(* Logix 5000 project; controller _GigaDiscovery vendor 1 type 14 code 244 rev 35.11; software revision 35.03; part 18 of 23 *)
(* tags used below, declared in another part *)
   Home_Timer : TIMER;
   Timer2 : TIMER;
   DC_Field_Motor_7 : UDT_CROUT;   // DC Field Motor 7 Gondola Contactor -Q16101E -Q16103E
   DC_Field_Pylon_Motors : UDT_CROUT;   // DC Field Pylon Motors Contactor -Q10101E -Q10103E
   FeedBack_Drives_Contactors : BOOL;
   Gate_Entry_Unlock_Selector : BOOL;   // -S30701F
   Gate_Exit_Unlock_Selector : BOOL;   // -S30705F
   Gate_Operator_Unlock_Selector : BOOL;   // -S30707F
   Gondola_Drive_Enable : UDT_CROUT;   // Gondola Drive Ch1-Ch2 Start Enable Contactors -Q16105E -Q16107E
   Gondola_Standstill_from_inertia : BOOL;
   I_Fbk_Platform_Main_Valve : UDT_DCS;   // Feedback Platform Main Valve -B21902I
   I_Fire_Interface : UDT_DCM;   // Page 44
   I_Gate_ENTER_G01_Closed : UDT_DCM;   // GATE ENTER (G01) -B25204I
   I_Gate_EXIT_G05_Closed : UDT_DCM;   // GATE EXIT (G05) -B25304I
   I_Gate_OPERATOR_Closed : UDT_DCM;   // GATE 4 OPERATOR RFID SENSOR - MOP -B25404J
   I_Gates_Closed : UDT_DCM;   // Gate Closed RFID series -B24802J
   I_GMB_RCC1_Temperature_OK : BOOL;   // +GMB_RCC1 Temperature OK -S40103E
   I_Gondola_Home_Position : BOOL;   // Gondola Home Position -B40002I -B40007I
   I_Gondola_Home_Position_Sensor_1 : UDT_DCM;   // Home Sensor Speed Check -B40002I
   I_Gondola_Home_Position_Sensor_2 : UDT_DCM;   // Home Sensor Speed Check -B40007I
   I_Platform_Closed : UDT_DCM;   // Platform Closed RFID Series -B22501J... -B22807J -B22801B
   I_Platform_Line_Min_Pressure_Switch : BOOL;   // Platform Line Minimum Pressure Switch -S21511B
   I_Platform_Line_Unlock_Pressure_Switch : BOOL;   // Unlock Platform Line Pressure Switch -S22006B
   I_Platform_Opened : UDT_DCM;   // Platform Opened RFID Series -Q23801J -Q23807J
   I_Platform_Pressure_on_Close_Circuit : BOOL;   // Platform Maximum Closing Pressure -S21510B
   I_Platform_Pressure_on_Open_Circuit : BOOL;   // Platform Maximum Opening Pressure -S21507B
   I_Pylon_Home_Ch1 : UDT_DCM;   // Home position Pylon Ch1 -B26002I
   I_Pylon_Home_Ch2 : UDT_DCM;   // Home position Pylon Ch2 -B26007I
   I_Pylon_Overlimit_Right : UDT_DCS;   // Pylon Overlimit Switchs -A26510I
   I_RCC_GSA_Temperature_OK : BOOL;   // +RCC_GSA Temperature OK -S50110G
   I_RCC_GSB_Temperature_OK : BOOL;   // +RCC_GSB Temperature OK -S52110G
   I_RCC_GSC_Temperature_OK : BOOL;   // +RCC_GSC Temperature OK -S54110G
   I_RCC_GSD_Temperature_OK : BOOL;   // +RCC_GSD Temperature OK -S56110G
   I_RCC_GSE_Temperature_OK : BOOL;   // +RCC_GSE Temperature OK -S58110G
   I_RCC_GSF_Temperature_OK : BOOL;   // +RCC_GSF Temperature OK -S60110G
   I_RCC_GSG_Temperature_OK : BOOL;   // +RCC_GSG Temperature OK -S62110G
   I_RCC_GSH_Temperature_OK : BOOL;   // +RCC_GSH Temperature OK -S64110G
   I_RESTRAINTS_Close_Limit_Switch : BOOL;   // Main Valve Close Limit Switch -B40508I
   I_RESTRAINTS_Open_Limit_Switch : BOOL;   // Main Valve Open Limit Switch -B40504I
   O_RESTRAINTS_Main_Valve : BOOL;   // Main Valve -B40501I
   O_RESTRAINTS_MainValve : UDT_CROUT;   // Main Valve -B40501I
   ONP : DINT;   // Optional Not Present
   Platform_Fbk_Valv_Close : BOOL;   // Platform Close Main Valve Limit Switch -B21909I
   Platform_Fbk_Valv_Open : BOOL;   // Platform Open Main Valve Limit Switch -B21905I
   Power_On_Delay : BOOL;
   Pylon_Contactor_OFF : BOOL;
   Pylon_Home_Position : UDT_DCM;   // Home position Pylon -B26002I -B26007I
   Pylon_Start_Drive_1_2 : UDT_CROUT;   // Pylon Start Drive 1 - 2 Contactors -Q9002H -Q9004H -Q10202G
   Pylon_Start_Drive_3_4 : UDT_CROUT;   // Pylon Start Drive 3 - 4 Contactors -Q9005H -Q9007H -Q12202G
   Pylon_Start_Drive_5_6 : UDT_CROUT;   // Pylon Start Drive 5 - 6 Contactors -Q9009E -Q9011E4 -Q14202G -Q14202G
   Pylon_Stopped_At_Home : BOOL;   // 5s
   Reset_Pulse : BOOL;
   RESTRAINTS_MainValve_PressTest : Valve_2_pos_monostable;
   RESTRAINTS_Rack : LapBar_Racks[41];
   RESTRAINTS_Sector : LapBars_Sector[9];
   RESTRAINTS_Unlock_Valve_Pressure : BOOL;
   Valves_Pressure_Discrepancy : DINT;
(* S_Input, continued *)

ROUTINE _04_Platform   (* ladder *)
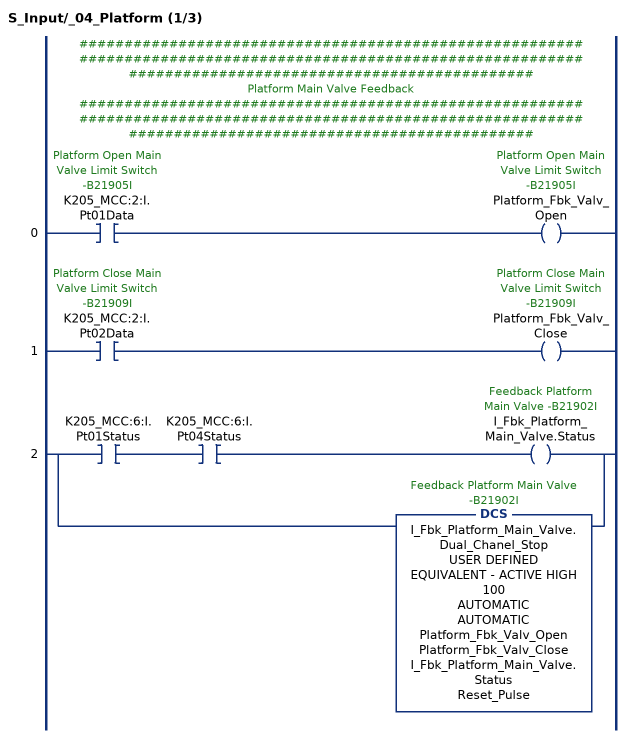
   // #############################################################################################################################################################
   // Platform Main Valve Feedback
   // #############################################################################################################################################################
   0: XIC(K205_MCC:2:I.Pt01Data)OTE(Platform_Fbk_Valv_Open);
   1: XIC(K205_MCC:2:I.Pt02Data)OTE(Platform_Fbk_Valv_Close);
   2: [XIC(K205_MCC:6:I.Pt01Status) XIC(K205_MCC:6:I.Pt04Status) OTE(I_Fbk_Platform_Main_Valve.Status) ,DCS(I_Fbk_Platform_Main_Valve.Dual_Chanel_Stop,USER DEFINED,EQUIVALENT - ACTIVE HIGH,100,AUTOMATIC,AUTOMATIC,Platform_Fbk_Valv_Open,Platform_Fbk_Valv_Close,I_Fbk_Platform_Main_Valve.Status,Reset_Pulse) ];
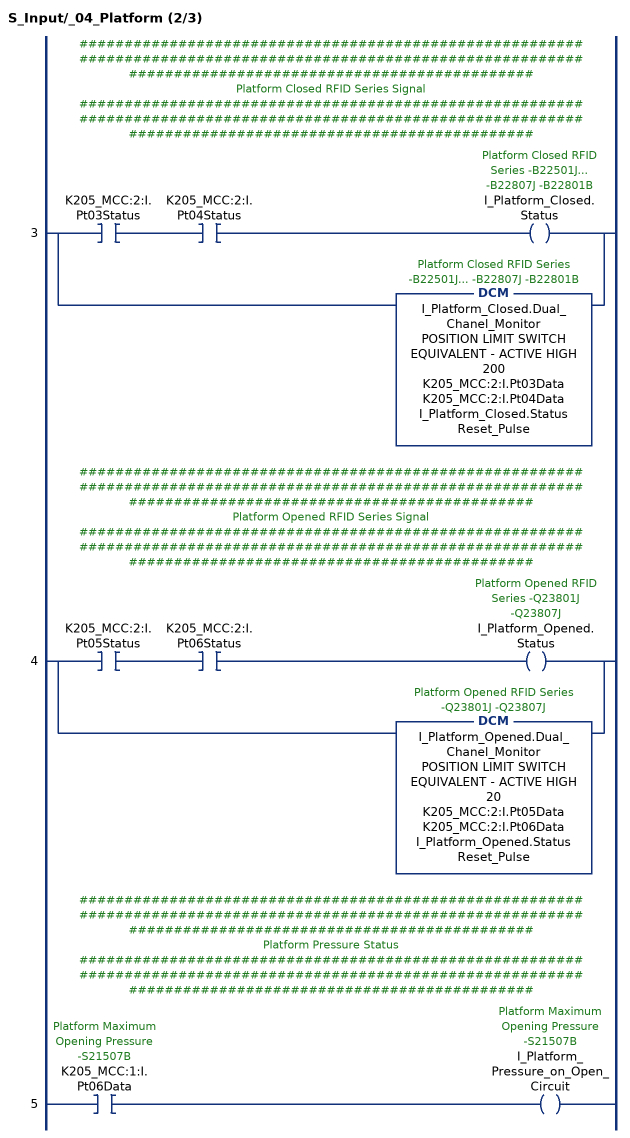
   // #############################################################################################################################################################
   // Platform Closed RFID Series Signal
   // #############################################################################################################################################################
   3: [XIC(K205_MCC:2:I.Pt03Status) XIC(K205_MCC:2:I.Pt04Status) OTE(I_Platform_Closed.Status) ,DCM(I_Platform_Closed.Dual_Chanel_Monitor,POSITION LIMIT SWITCH,EQUIVALENT - ACTIVE HIGH,200,K205_MCC:2:I.Pt03Data,K205_MCC:2:I.Pt04Data,I_Platform_Closed.Status,Reset_Pulse) ];
   // #############################################################################################################################################################
   // Platform Opened RFID Series Signal
   // #############################################################################################################################################################
   4: [XIC(K205_MCC:2:I.Pt05Status) XIC(K205_MCC:2:I.Pt06Status) OTE(I_Platform_Opened.Status) ,DCM(I_Platform_Opened.Dual_Chanel_Monitor,POSITION LIMIT SWITCH,EQUIVALENT - ACTIVE HIGH,20,K205_MCC:2:I.Pt05Data,K205_MCC:2:I.Pt06Data,I_Platform_Opened.Status,Reset_Pulse) ];
   // #############################################################################################################################################################
   // Platform Pressure Status
   // #############################################################################################################################################################
   5: XIC(K205_MCC:1:I.Pt06Data)OTE(I_Platform_Pressure_on_Open_Circuit);
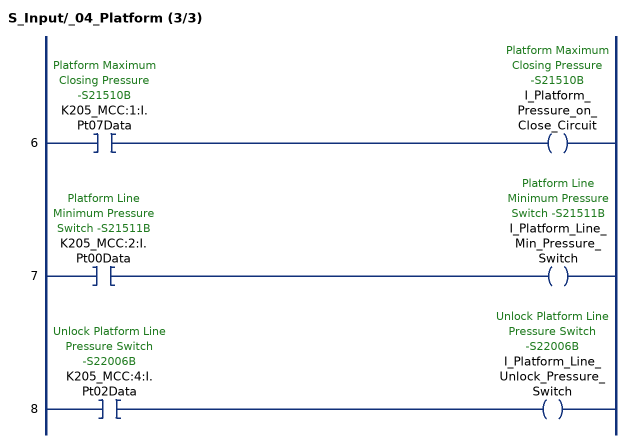
   6: XIC(K205_MCC:1:I.Pt07Data)OTE(I_Platform_Pressure_on_Close_Circuit);
   7: XIC(K205_MCC:2:I.Pt00Data)OTE(I_Platform_Line_Min_Pressure_Switch);
   8: XIC(K205_MCC:4:I.Pt02Data)OTE(I_Platform_Line_Unlock_Pressure_Switch);
END_ROUTINE

ROUTINE _05_Pylon   (* ladder *)
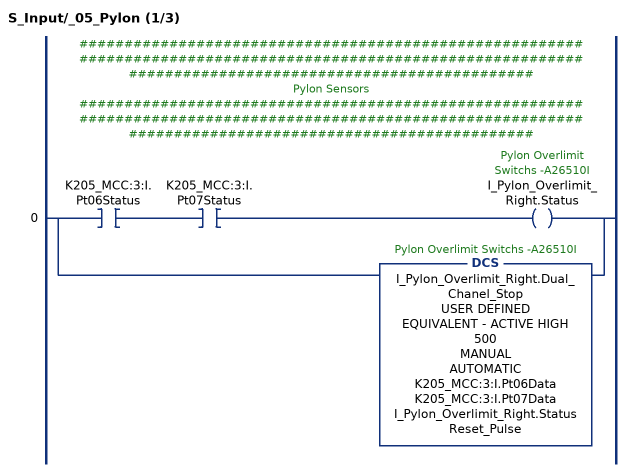
   // #############################################################################################################################################################
   // Pylon Sensors
   // #############################################################################################################################################################
   0: [XIC(K205_MCC:3:I.Pt06Status) XIC(K205_MCC:3:I.Pt07Status) OTE(I_Pylon_Overlimit_Right.Status) ,DCS(I_Pylon_Overlimit_Right.Dual_Chanel_Stop,USER DEFINED,EQUIVALENT - ACTIVE HIGH,500,MANUAL,AUTOMATIC,K205_MCC:3:I.Pt06Data,K205_MCC:3:I.Pt07Data,I_Pylon_Overlimit_Right.Status,Reset_Pulse) ];
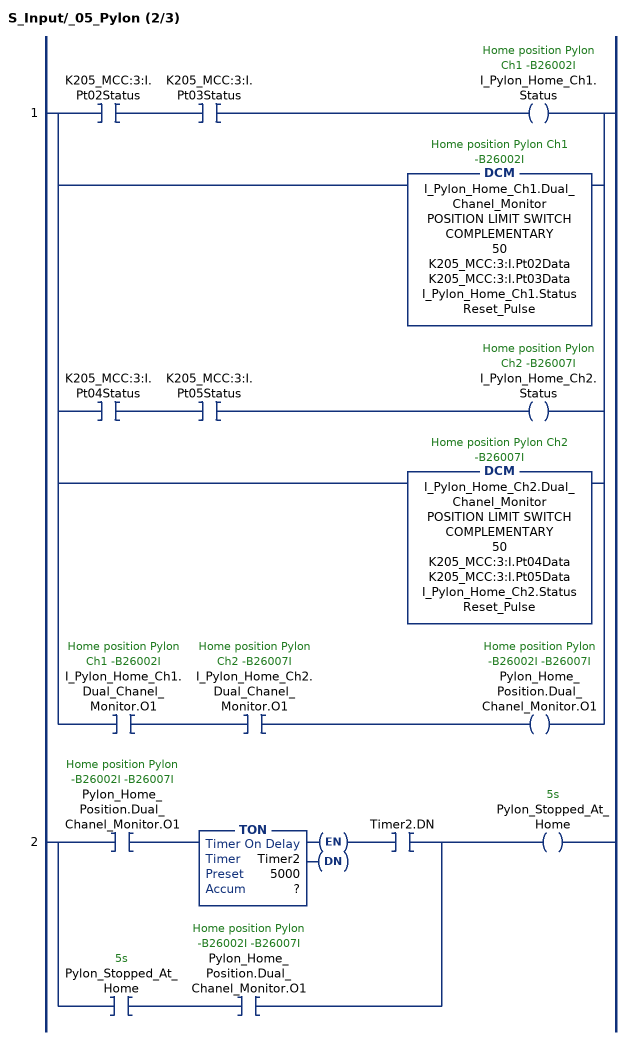
   1: [[XIC(K205_MCC:3:I.Pt02Status) XIC(K205_MCC:3:I.Pt03Status) OTE(I_Pylon_Home_Ch1.Status) ,DCM(I_Pylon_Home_Ch1.Dual_Chanel_Monitor,POSITION LIMIT SWITCH,COMPLEMENTARY,50,K205_MCC:3:I.Pt02Data,K205_MCC:3:I.Pt03Data,I_Pylon_Home_Ch1.Status,Reset_Pulse) ] ,[XIC(K205_MCC:3:I.Pt04Status) XIC(K205_MCC:3:I.Pt05Status) OTE(I_Pylon_Home_Ch2.Status) ,DCM(I_Pylon_Home_Ch2.Dual_Chanel_Monitor,POSITION LIMIT SWITCH,COMPLEMENTARY,50,K205_MCC:3:I.Pt04Data,K205_MCC:3:I.Pt05Data,I_Pylon_Home_Ch2.Status,Reset_Pulse) ] ,XIC(I_Pylon_Home_Ch1.Dual_Chanel_Monitor.O1) XIC(I_Pylon_Home_Ch2.Dual_Chanel_Monitor.O1) OTE(Pylon_Home_Position.Dual_Chanel_Monitor.O1) ];
   2: [XIC(Pylon_Home_Position.Dual_Chanel_Monitor.O1) TON(Timer2,?,?) XIC(Timer2.DN) ,XIC(Pylon_Stopped_At_Home) XIC(Pylon_Home_Position.Dual_Chanel_Monitor.O1) ]OTE(Pylon_Stopped_At_Home);
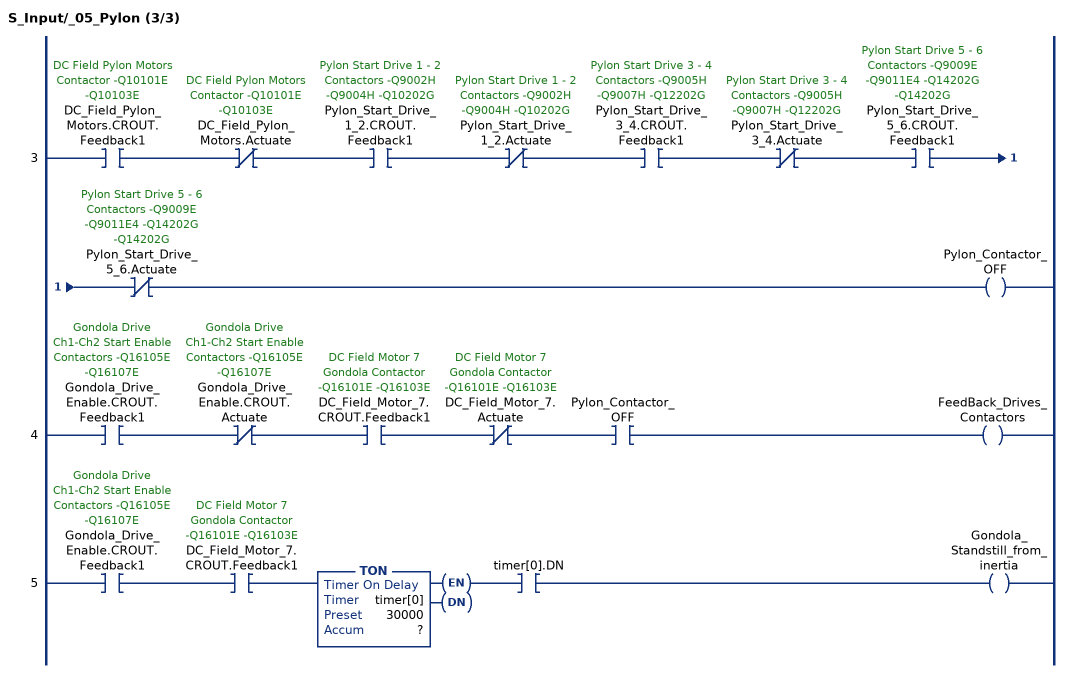
   3: XIC(DC_Field_Pylon_Motors.CROUT.Feedback1)XIO(DC_Field_Pylon_Motors.Actuate)XIC(Pylon_Start_Drive_1_2.CROUT.Feedback1)XIO(Pylon_Start_Drive_1_2.Actuate)XIC(Pylon_Start_Drive_3_4.CROUT.Feedback1)XIO(Pylon_Start_Drive_3_4.Actuate)XIC(Pylon_Start_Drive_5_6.CROUT.Feedback1)XIO(Pylon_Start_Drive_5_6.Actuate)OTE(Pylon_Contactor_OFF);
   4: XIC(Gondola_Drive_Enable.CROUT.Feedback1)XIO(Gondola_Drive_Enable.CROUT.Actuate)XIC(DC_Field_Motor_7.CROUT.Feedback1)XIO(DC_Field_Motor_7.Actuate)XIC(Pylon_Contactor_OFF)OTE(FeedBack_Drives_Contactors);
   5: XIC(Gondola_Drive_Enable.CROUT.Feedback1)XIC(DC_Field_Motor_7.CROUT.Feedback1)TON(timer[0],?,?)XIC(timer[0].DN)OTE(Gondola_Standstill_from_inertia);
END_ROUTINE

ROUTINE _06_RCC   (* ladder *)
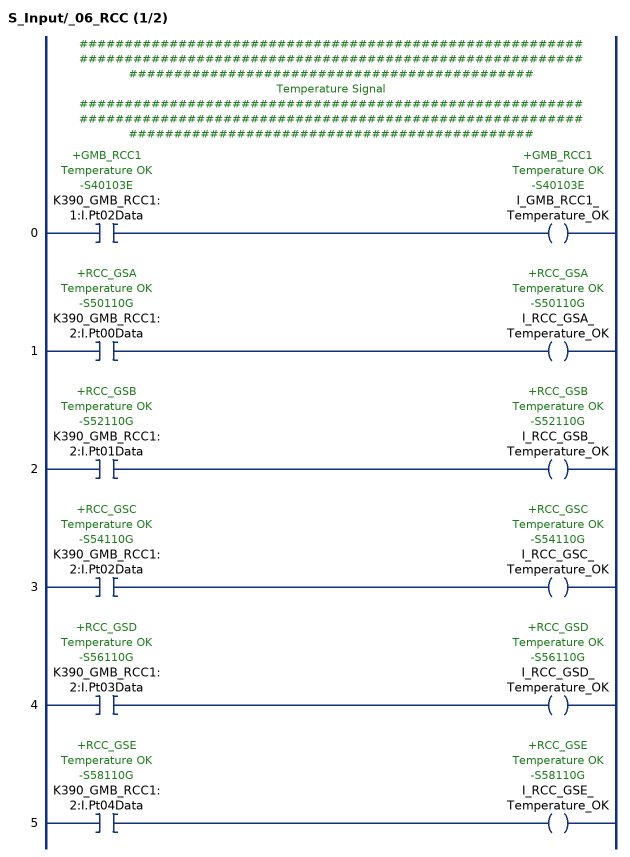
   // #############################################################################################################################################################
   //   Temperature Signal
   // #############################################################################################################################################################
   0: XIC(K390_GMB_RCC1:1:I.Pt02Data)OTE(I_GMB_RCC1_Temperature_OK);
   1: XIC(K390_GMB_RCC1:2:I.Pt00Data)OTE(I_RCC_GSA_Temperature_OK);
   2: XIC(K390_GMB_RCC1:2:I.Pt01Data)OTE(I_RCC_GSB_Temperature_OK);
   3: XIC(K390_GMB_RCC1:2:I.Pt02Data)OTE(I_RCC_GSC_Temperature_OK);
   4: XIC(K390_GMB_RCC1:2:I.Pt03Data)OTE(I_RCC_GSD_Temperature_OK);
   5: XIC(K390_GMB_RCC1:2:I.Pt04Data)OTE(I_RCC_GSE_Temperature_OK);
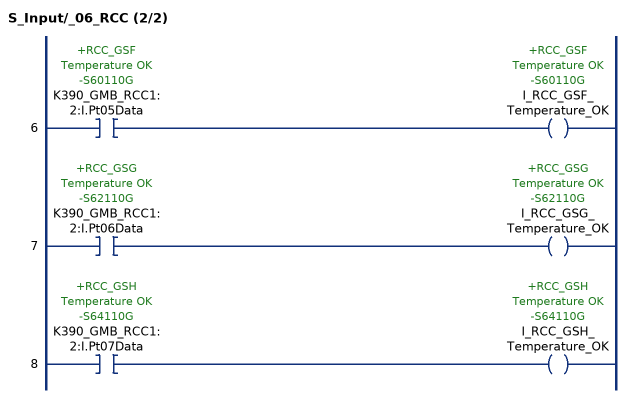
   6: XIC(K390_GMB_RCC1:2:I.Pt05Data)OTE(I_RCC_GSF_Temperature_OK);
   7: XIC(K390_GMB_RCC1:2:I.Pt06Data)OTE(I_RCC_GSG_Temperature_OK);
   8: XIC(K390_GMB_RCC1:2:I.Pt07Data)OTE(I_RCC_GSH_Temperature_OK);
END_ROUTINE

ROUTINE _07_Gate   (* ladder *)
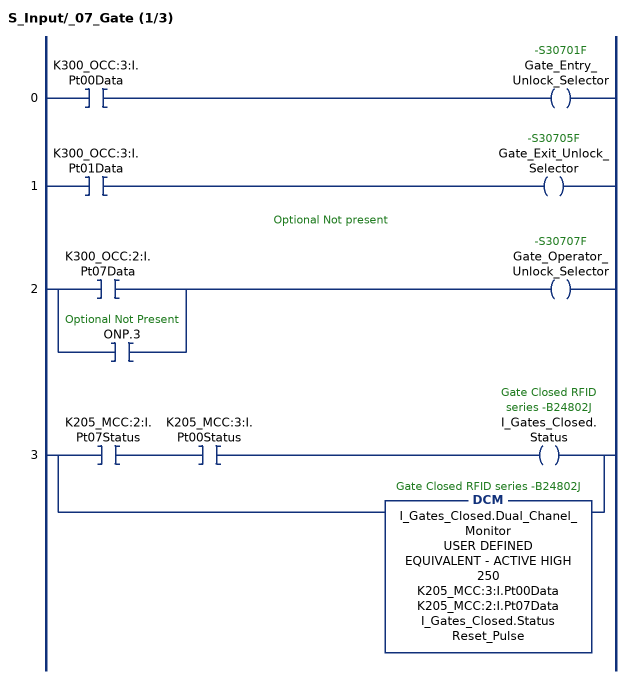
   0: XIC(K300_OCC:3:I.Pt00Data)OTE(Gate_Entry_Unlock_Selector);
   1: XIC(K300_OCC:3:I.Pt01Data)OTE(Gate_Exit_Unlock_Selector);
   // Optional Not present
   2: [XIC(K300_OCC:2:I.Pt07Data) ,XIC(ONP.3) ]OTE(Gate_Operator_Unlock_Selector);
   3: [XIC(K205_MCC:2:I.Pt07Status) XIC(K205_MCC:3:I.Pt00Status) OTE(I_Gates_Closed.Status) ,DCM(I_Gates_Closed.Dual_Chanel_Monitor,USER DEFINED,EQUIVALENT - ACTIVE HIGH,250,K205_MCC:3:I.Pt00Data,K205_MCC:2:I.Pt07Data,I_Gates_Closed.Status,Reset_Pulse) ];
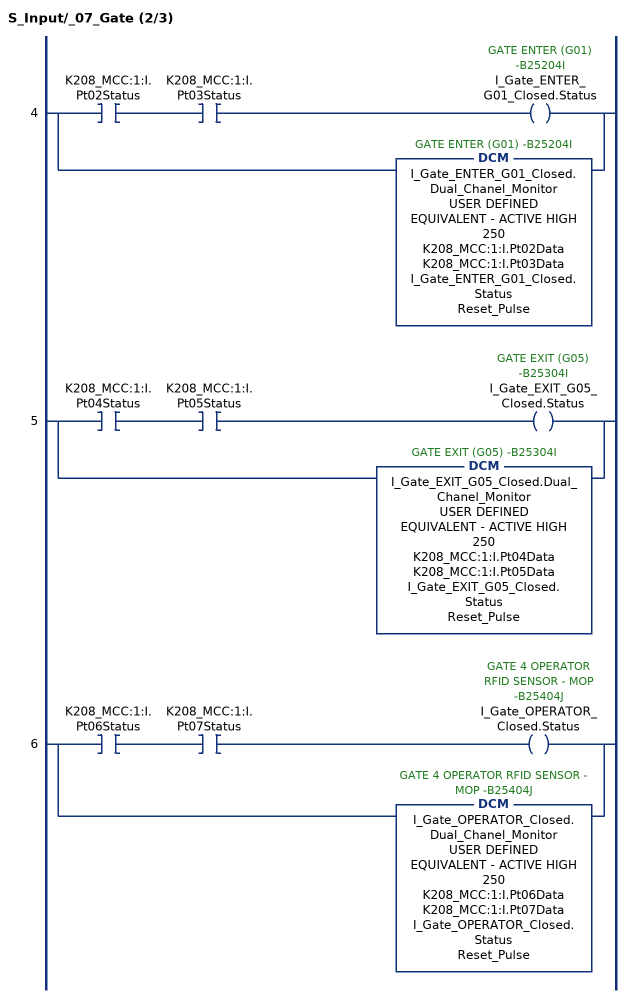
   4: [XIC(K208_MCC:1:I.Pt02Status) XIC(K208_MCC:1:I.Pt03Status) OTE(I_Gate_ENTER_G01_Closed.Status) ,DCM(I_Gate_ENTER_G01_Closed.Dual_Chanel_Monitor,USER DEFINED,EQUIVALENT - ACTIVE HIGH,250,K208_MCC:1:I.Pt02Data,K208_MCC:1:I.Pt03Data,I_Gate_ENTER_G01_Closed.Status,Reset_Pulse) ];
   5: [XIC(K208_MCC:1:I.Pt04Status) XIC(K208_MCC:1:I.Pt05Status) OTE(I_Gate_EXIT_G05_Closed.Status) ,DCM(I_Gate_EXIT_G05_Closed.Dual_Chanel_Monitor,USER DEFINED,EQUIVALENT - ACTIVE HIGH,250,K208_MCC:1:I.Pt04Data,K208_MCC:1:I.Pt05Data,I_Gate_EXIT_G05_Closed.Status,Reset_Pulse) ];
   6: [XIC(K208_MCC:1:I.Pt06Status) XIC(K208_MCC:1:I.Pt07Status) OTE(I_Gate_OPERATOR_Closed.Status) ,DCM(I_Gate_OPERATOR_Closed.Dual_Chanel_Monitor,USER DEFINED,EQUIVALENT - ACTIVE HIGH,250,K208_MCC:1:I.Pt06Data,K208_MCC:1:I.Pt07Data,I_Gate_OPERATOR_Closed.Status,Reset_Pulse) ];
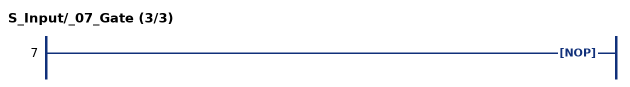
   7: NOP();
END_ROUTINE

ROUTINE _08_Gondola   (* ladder *)
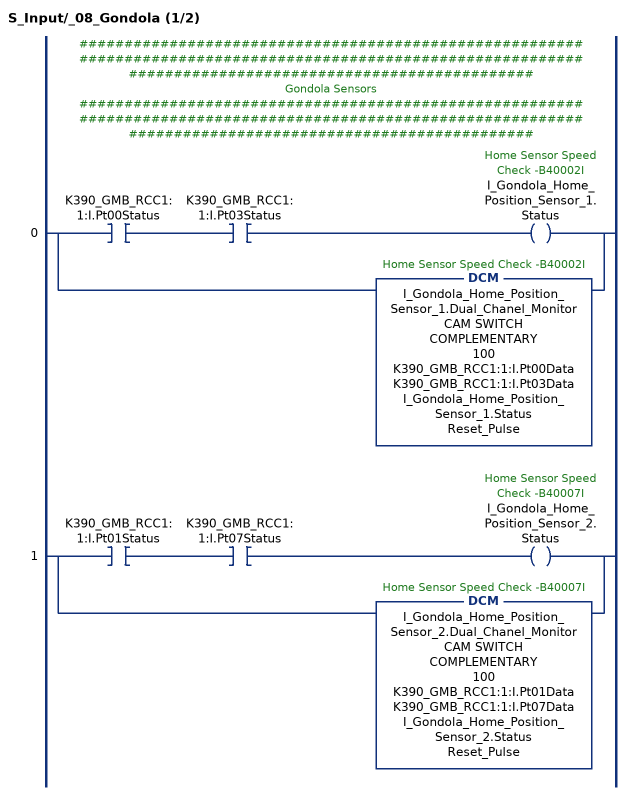
   // #############################################################################################################################################################
   // Gondola Sensors
   // #############################################################################################################################################################
   0: [XIC(K390_GMB_RCC1:1:I.Pt00Status) XIC(K390_GMB_RCC1:1:I.Pt03Status) OTE(I_Gondola_Home_Position_Sensor_1.Status) ,DCM(I_Gondola_Home_Position_Sensor_1.Dual_Chanel_Monitor,CAM SWITCH,COMPLEMENTARY,100,K390_GMB_RCC1:1:I.Pt00Data,K390_GMB_RCC1:1:I.Pt03Data,I_Gondola_Home_Position_Sensor_1.Status,Reset_Pulse) ];
   1: [XIC(K390_GMB_RCC1:1:I.Pt01Status) XIC(K390_GMB_RCC1:1:I.Pt07Status) OTE(I_Gondola_Home_Position_Sensor_2.Status) ,DCM(I_Gondola_Home_Position_Sensor_2.Dual_Chanel_Monitor,CAM SWITCH,COMPLEMENTARY,100,K390_GMB_RCC1:1:I.Pt01Data,K390_GMB_RCC1:1:I.Pt07Data,I_Gondola_Home_Position_Sensor_2.Status,Reset_Pulse) ];
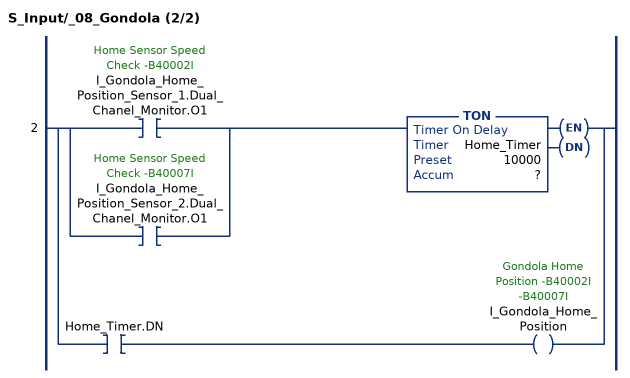
   2: [[XIC(I_Gondola_Home_Position_Sensor_1.Dual_Chanel_Monitor.O1) ,XIC(I_Gondola_Home_Position_Sensor_2.Dual_Chanel_Monitor.O1) ] TON(Home_Timer,?,?) ,XIC(Home_Timer.DN) OTE(I_Gondola_Home_Position) ];
END_ROUTINE

ROUTINE _09_External_Interface   (* ladder *)
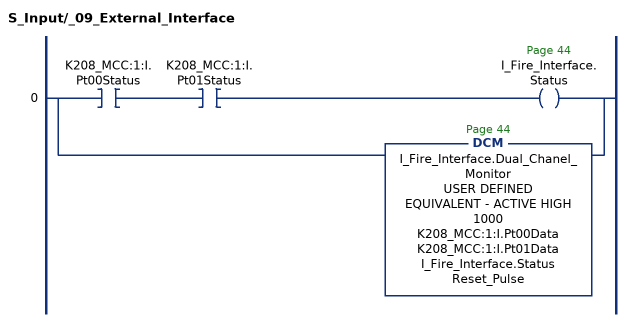
   0: [XIC(K208_MCC:1:I.Pt00Status) XIC(K208_MCC:1:I.Pt01Status) OTE(I_Fire_Interface.Status) ,DCM(I_Fire_Interface.Dual_Chanel_Monitor,USER DEFINED,EQUIVALENT - ACTIVE HIGH,1000,K208_MCC:1:I.Pt00Data,K208_MCC:1:I.Pt01Data,I_Fire_Interface.Status,Reset_Pulse) ];
END_ROUTINE

ROUTINE Main   (* ladder *)
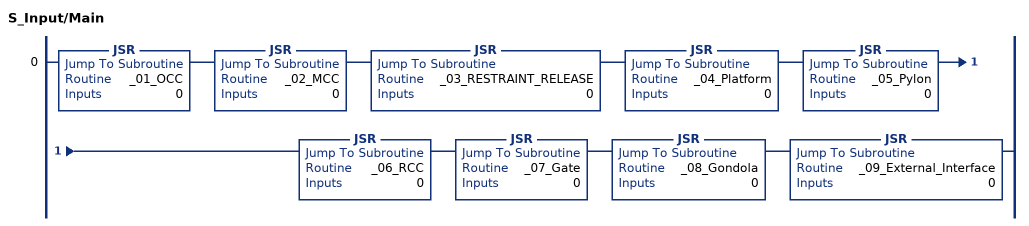
   0: JSR(_01_OCC,0)JSR(_02_MCC,0)JSR(_03_RESTRAINT_RELEASE,0)JSR(_04_Platform,0)JSR(_05_Pylon,0)JSR(_06_RCC,0)JSR(_07_Gate,0)JSR(_08_Gondola,0)JSR(_09_External_Interface,0);
END_ROUTINE
END_PROGRAM

PROGRAM S_Output   (* main routine Main, safety *)
VAR
   Os : DINT;
   Timer : TIMER[10] := ([0].PRE := 1200000, [0].EN := 1, [0].DN := 1, [1].PRE := 5000, [2].PRE := 20000, [2].ACC := 20000, [3].PRE := 1200000, [3].ACC := 1200000);
END_VAR

ROUTINE _02_Lap_Bars   (* ladder *)
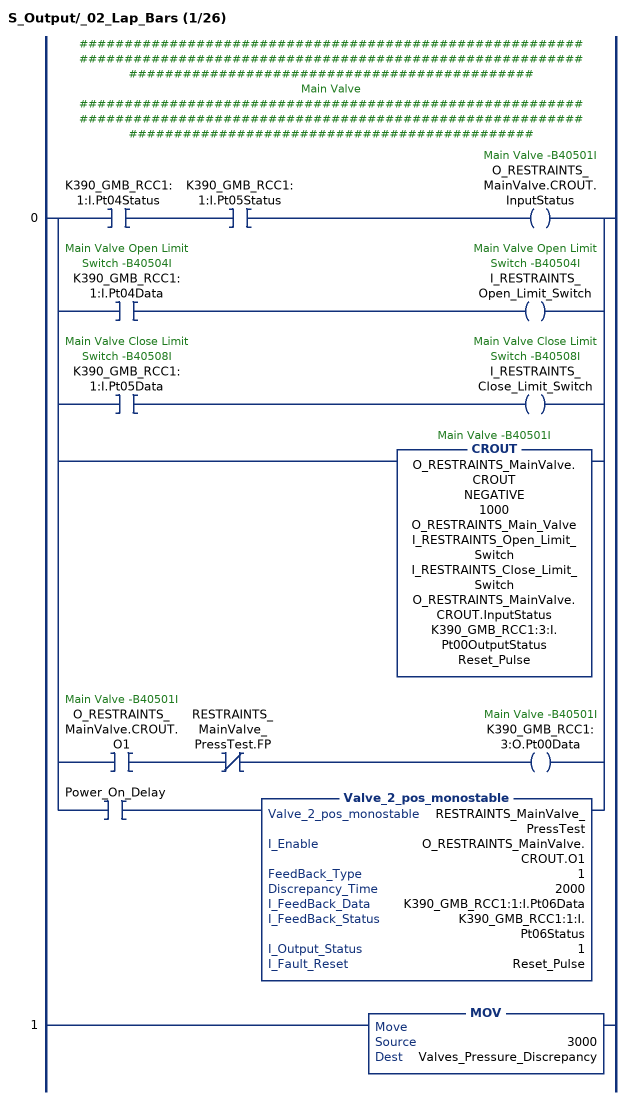
   // #############################################################################################################################################################
   // Main Valve
   // #############################################################################################################################################################
   0: [XIC(K390_GMB_RCC1:1:I.Pt04Status) XIC(K390_GMB_RCC1:1:I.Pt05Status) OTE(O_RESTRAINTS_MainValve.CROUT.InputStatus) ,XIC(K390_GMB_RCC1:1:I.Pt04Data) OTE(I_RESTRAINTS_Open_Limit_Switch) ,XIC(K390_GMB_RCC1:1:I.Pt05Data) OTE(I_RESTRAINTS_Close_Limit_Switch) ,CROUT(O_RESTRAINTS_MainValve.CROUT,NEGATIVE,1000,O_RESTRAINTS_Main_Valve,I_RESTRAINTS_Open_Limit_Switch,I_RESTRAINTS_Close_Limit_Switch,O_RESTRAINTS_MainValve.CROUT.InputStatus,K390_GMB_RCC1:3:I.Pt00OutputStatus,Reset_Pulse) ,XIC(O_RESTRAINTS_MainValve.CROUT.O1) XIO(RESTRAINTS_MainValve_PressTest.FP) OTE(K390_GMB_RCC1:3:O.Pt00Data) ,XIC(Power_On_Delay) Valve_2_pos_monostable(RESTRAINTS_MainValve_PressTest,O_RESTRAINTS_MainValve.CROUT.O1,1,2000,K390_GMB_RCC1:1:I.Pt06Data,K390_GMB_RCC1:1:I.Pt06Status,1,Reset_Pulse) ];
   1: MOV(3000,Valves_Pressure_Discrepancy);
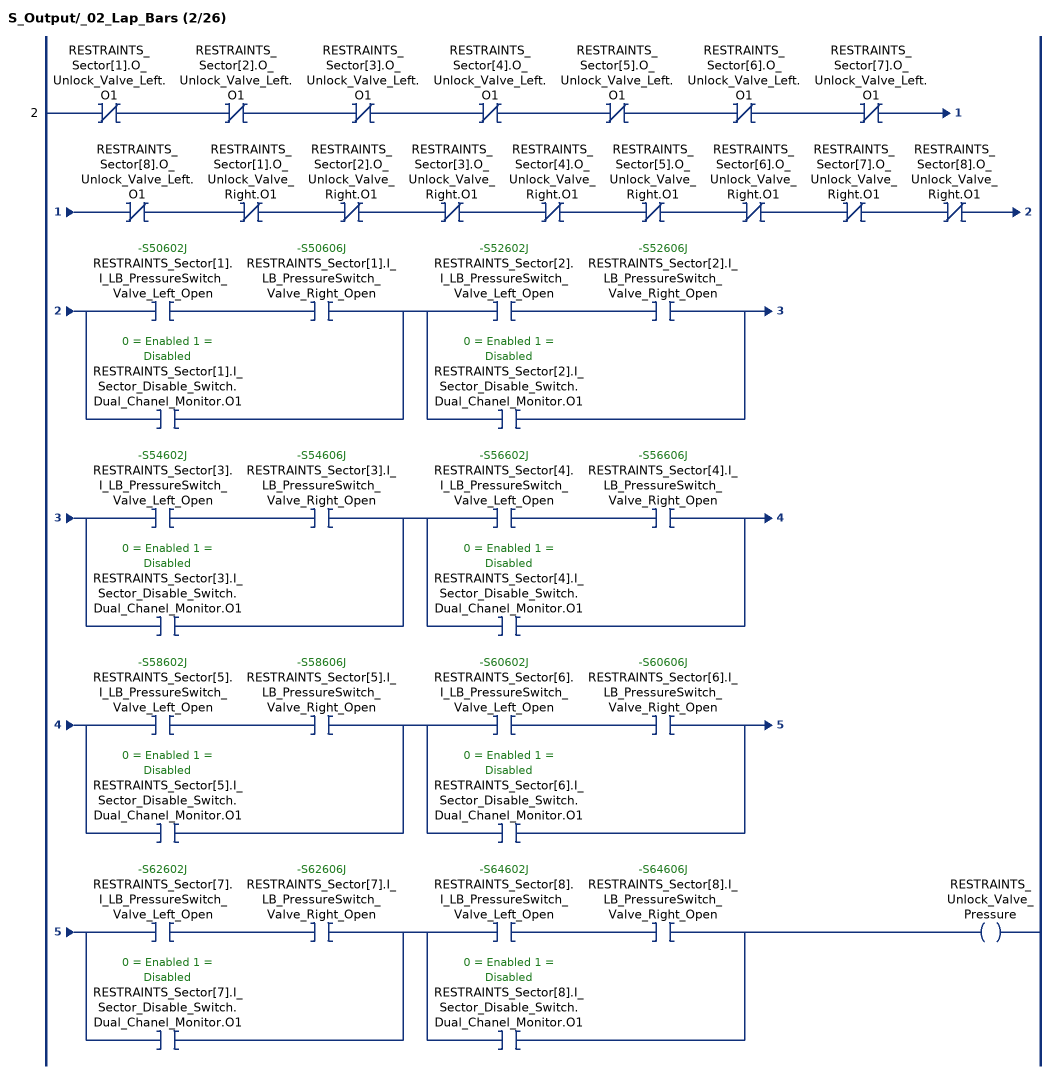
   2: XIO(RESTRAINTS_Sector[1].O_Unlock_Valve_Left.O1)XIO(RESTRAINTS_Sector[2].O_Unlock_Valve_Left.O1)XIO(RESTRAINTS_Sector[3].O_Unlock_Valve_Left.O1)XIO(RESTRAINTS_Sector[4].O_Unlock_Valve_Left.O1)XIO(RESTRAINTS_Sector[5].O_Unlock_Valve_Left.O1)XIO(RESTRAINTS_Sector[6].O_Unlock_Valve_Left.O1)XIO(RESTRAINTS_Sector[7].O_Unlock_Valve_Left.O1)XIO(RESTRAINTS_Sector[8].O_Unlock_Valve_Left.O1)XIO(RESTRAINTS_Sector[1].O_Unlock_Valve_Right.O1)XIO(RESTRAINTS_Sector[2].O_Unlock_Valve_Right.O1)XIO(RESTRAINTS_Sector[3].O_Unlock_Valve_Right.O1)XIO(RESTRAINTS_Sector[4].O_Unlock_Valve_Right.O1)XIO(RESTRAINTS_Sector[5].O_Unlock_Valve_Right.O1)XIO(RESTRAINTS_Sector[6].O_Unlock_Valve_Right.O1)XIO(RESTRAINTS_Sector[7].O_Unlock_Valve_Right.O1)XIO(RESTRAINTS_Sector[8].O_Unlock_Valve_Right.O1)[XIC(RESTRAINTS_Sector[1].I_LB_PressureSwitch_Valve_Left_Open) XIC(RESTRAINTS_Sector[1].I_LB_PressureSwitch_Valve_Right_Open) ,XIC(RESTRAINTS_Sector[1].I_Sector_Disable_Switch.Dual_Chanel_Monitor.O1) ][XIC(RESTRAINTS_Sector[2].I_LB_PressureSwitch_Valve_Left_Open) XIC(RESTRAINTS_Sector[2].I_LB_PressureSwitch_Valve_Right_Open) ,XIC(RESTRAINTS_Sector[2].I_Sector_Disable_Switch.Dual_Chanel_Monitor.O1) ][XIC(RESTRAINTS_Sector[3].I_LB_PressureSwitch_Valve_Left_Open) XIC(RESTRAINTS_Sector[3].I_LB_PressureSwitch_Valve_Right_Open) ,XIC(RESTRAINTS_Sector[3].I_Sector_Disable_Switch.Dual_Chanel_Monitor.O1) ][XIC(RESTRAINTS_Sector[4].I_LB_PressureSwitch_Valve_Left_Open) XIC(RESTRAINTS_Sector[4].I_LB_PressureSwitch_Valve_Right_Open) ,XIC(RESTRAINTS_Sector[4].I_Sector_Disable_Switch.Dual_Chanel_Monitor.O1) ][XIC(RESTRAINTS_Sector[5].I_LB_PressureSwitch_Valve_Left_Open) XIC(RESTRAINTS_Sector[5].I_LB_PressureSwitch_Valve_Right_Open) ,XIC(RESTRAINTS_Sector[5].I_Sector_Disable_Switch.Dual_Chanel_Monitor.O1) ][XIC(RESTRAINTS_Sector[6].I_LB_PressureSwitch_Valve_Left_Open) XIC(RESTRAINTS_Sector[6].I_LB_PressureSwitch_Valve_Right_Open) ,XIC(RESTRAINTS_Sector[6].I_Sector_Disable_Switch.Dual_Chanel_Monitor.O1) ][XIC(RESTRAINTS_Sector[7].I_LB_PressureSwitch_Valve_Left_Open) XIC(RESTRAINTS_Sector[7].I_LB_PressureSwitch_Valve_Right_Open) ,XIC(RESTRAINTS_Sector[7].I_Sector_Disable_Switch.Dual_Chanel_Monitor.O1) ][XIC(RESTRAINTS_Sector[8].I_LB_PressureSwitch_Valve_Left_Open) XIC(RESTRAINTS_Sector[8].I_LB_PressureSwitch_Valve_Right_Open) ,XIC(RESTRAINTS_Sector[8].I_Sector_Disable_Switch.Dual_Chanel_Monitor.O1) ]OTE(RESTRAINTS_Unlock_Valve_Pressure);
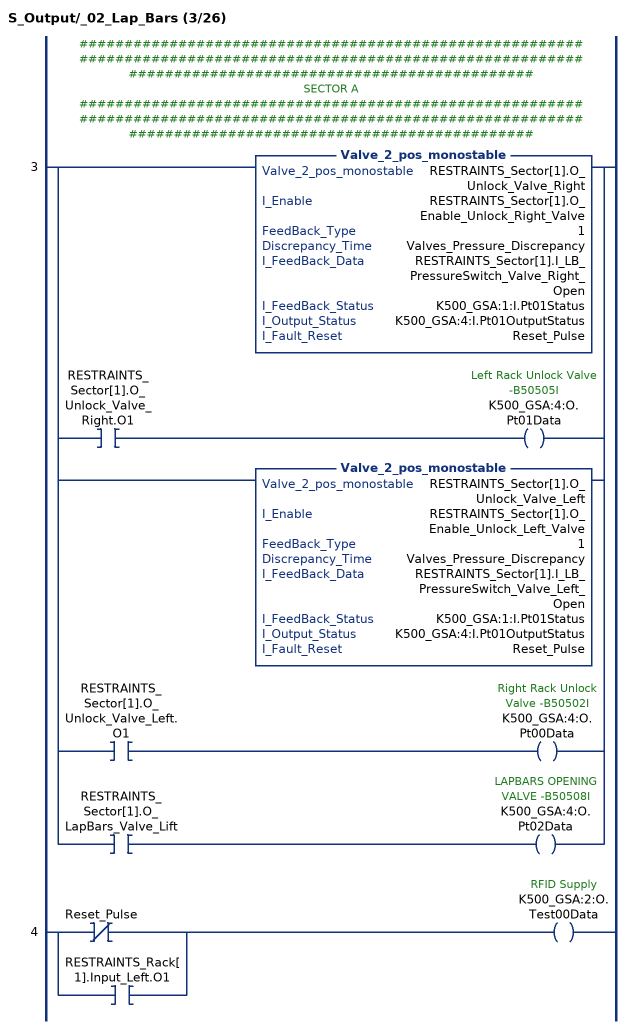
   // #############################################################################################################################################################
   // SECTOR A
   // #############################################################################################################################################################
   3: [[Valve_2_pos_monostable(RESTRAINTS_Sector[1].O_Unlock_Valve_Right,RESTRAINTS_Sector[1].O_Enable_Unlock_Right_Valve,1,Valves_Pressure_Discrepancy,RESTRAINTS_Sector[1].I_LB_PressureSwitch_Valve_Right_Open,K500_GSA:1:I.Pt01Status,K500_GSA:4:I.Pt01OutputStatus,Reset_Pulse) ,XIC(RESTRAINTS_Sector[1].O_Unlock_Valve_Right.O1) OTE(K500_GSA:4:O.Pt01Data) ] ,[Valve_2_pos_monostable(RESTRAINTS_Sector[1].O_Unlock_Valve_Left,RESTRAINTS_Sector[1].O_Enable_Unlock_Left_Valve,1,Valves_Pressure_Discrepancy,RESTRAINTS_Sector[1].I_LB_PressureSwitch_Valve_Left_Open,K500_GSA:1:I.Pt01Status,K500_GSA:4:I.Pt01OutputStatus,Reset_Pulse) ,XIC(RESTRAINTS_Sector[1].O_Unlock_Valve_Left.O1) OTE(K500_GSA:4:O.Pt00Data) ] ,XIC(RESTRAINTS_Sector[1].O_LapBars_Valve_Lift) OTE(K500_GSA:4:O.Pt02Data) ];
   4: [XIO(Reset_Pulse) ,XIC(RESTRAINTS_Rack[1].Input_Left.O1) ]OTE(K500_GSA:2:O.Test00Data);
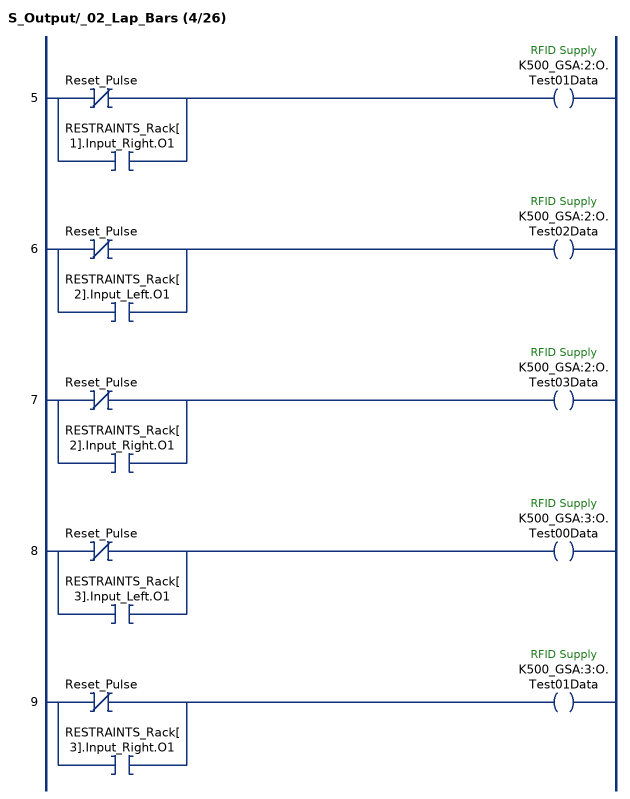
   5: [XIO(Reset_Pulse) ,XIC(RESTRAINTS_Rack[1].Input_Right.O1) ]OTE(K500_GSA:2:O.Test01Data);
   6: [XIO(Reset_Pulse) ,XIC(RESTRAINTS_Rack[2].Input_Left.O1) ]OTE(K500_GSA:2:O.Test02Data);
   7: [XIO(Reset_Pulse) ,XIC(RESTRAINTS_Rack[2].Input_Right.O1) ]OTE(K500_GSA:2:O.Test03Data);
   8: [XIO(Reset_Pulse) ,XIC(RESTRAINTS_Rack[3].Input_Left.O1) ]OTE(K500_GSA:3:O.Test00Data);
   9: [XIO(Reset_Pulse) ,XIC(RESTRAINTS_Rack[3].Input_Right.O1) ]OTE(K500_GSA:3:O.Test01Data);
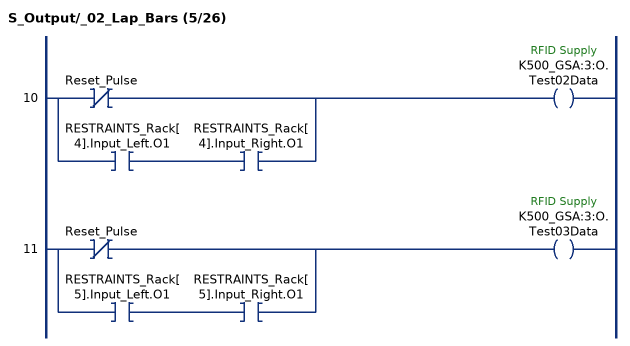
   10: [XIO(Reset_Pulse) ,XIC(RESTRAINTS_Rack[4].Input_Left.O1) XIC(RESTRAINTS_Rack[4].Input_Right.O1) ]OTE(K500_GSA:3:O.Test02Data);
   11: [XIO(Reset_Pulse) ,XIC(RESTRAINTS_Rack[5].Input_Left.O1) XIC(RESTRAINTS_Rack[5].Input_Right.O1) ]OTE(K500_GSA:3:O.Test03Data);
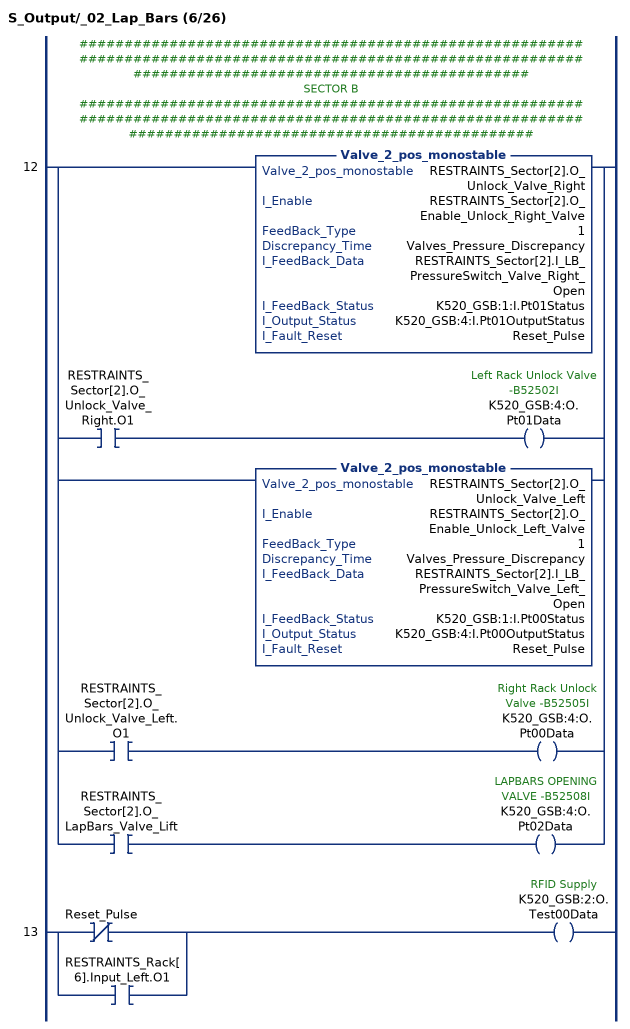
   // ############################################################################################################################################################
   // SECTOR B
   // #############################################################################################################################################################
   12: [[Valve_2_pos_monostable(RESTRAINTS_Sector[2].O_Unlock_Valve_Right,RESTRAINTS_Sector[2].O_Enable_Unlock_Right_Valve,1,Valves_Pressure_Discrepancy,RESTRAINTS_Sector[2].I_LB_PressureSwitch_Valve_Right_Open,K520_GSB:1:I.Pt01Status,K520_GSB:4:I.Pt01OutputStatus,Reset_Pulse) ,XIC(RESTRAINTS_Sector[2].O_Unlock_Valve_Right.O1) OTE(K520_GSB:4:O.Pt01Data) ] ,[Valve_2_pos_monostable(RESTRAINTS_Sector[2].O_Unlock_Valve_Left,RESTRAINTS_Sector[2].O_Enable_Unlock_Left_Valve,1,Valves_Pressure_Discrepancy,RESTRAINTS_Sector[2].I_LB_PressureSwitch_Valve_Left_Open,K520_GSB:1:I.Pt00Status,K520_GSB:4:I.Pt00OutputStatus,Reset_Pulse) ,XIC(RESTRAINTS_Sector[2].O_Unlock_Valve_Left.O1) OTE(K520_GSB:4:O.Pt00Data) ] ,XIC(RESTRAINTS_Sector[2].O_LapBars_Valve_Lift) OTE(K520_GSB:4:O.Pt02Data) ];
   13: [XIO(Reset_Pulse) ,XIC(RESTRAINTS_Rack[6].Input_Left.O1) ]OTE(K520_GSB:2:O.Test00Data);
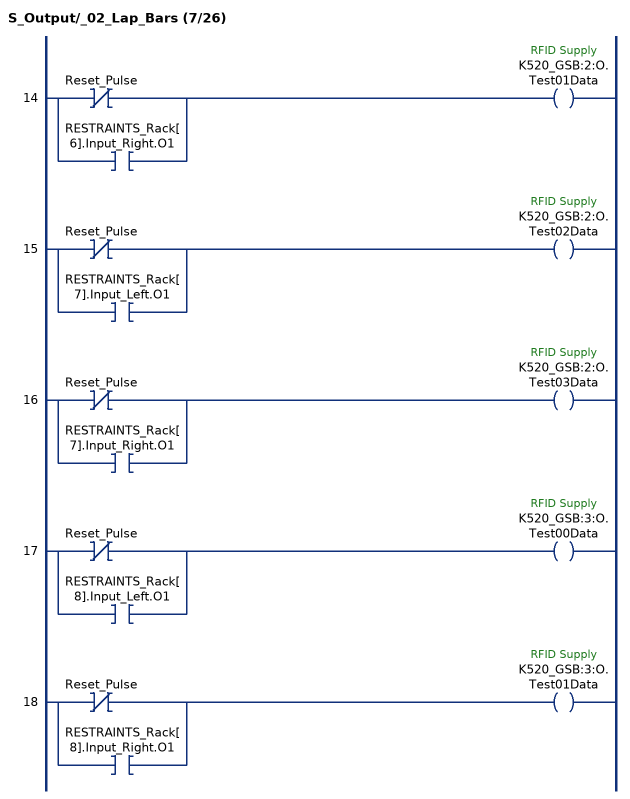
   14: [XIO(Reset_Pulse) ,XIC(RESTRAINTS_Rack[6].Input_Right.O1) ]OTE(K520_GSB:2:O.Test01Data);
   15: [XIO(Reset_Pulse) ,XIC(RESTRAINTS_Rack[7].Input_Left.O1) ]OTE(K520_GSB:2:O.Test02Data);
   16: [XIO(Reset_Pulse) ,XIC(RESTRAINTS_Rack[7].Input_Right.O1) ]OTE(K520_GSB:2:O.Test03Data);
   17: [XIO(Reset_Pulse) ,XIC(RESTRAINTS_Rack[8].Input_Left.O1) ]OTE(K520_GSB:3:O.Test00Data);
   18: [XIO(Reset_Pulse) ,XIC(RESTRAINTS_Rack[8].Input_Right.O1) ]OTE(K520_GSB:3:O.Test01Data);
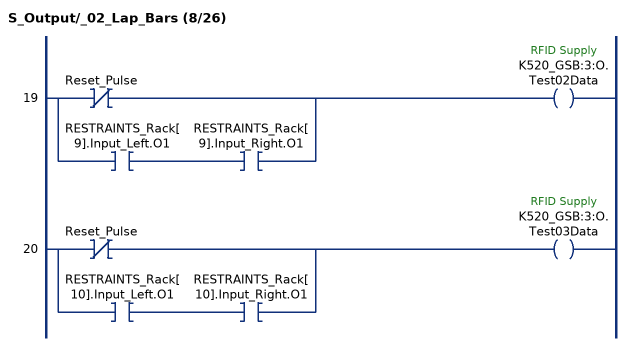
   19: [XIO(Reset_Pulse) ,XIC(RESTRAINTS_Rack[9].Input_Left.O1) XIC(RESTRAINTS_Rack[9].Input_Right.O1) ]OTE(K520_GSB:3:O.Test02Data);
   20: [XIO(Reset_Pulse) ,XIC(RESTRAINTS_Rack[10].Input_Left.O1) XIC(RESTRAINTS_Rack[10].Input_Right.O1) ]OTE(K520_GSB:3:O.Test03Data);
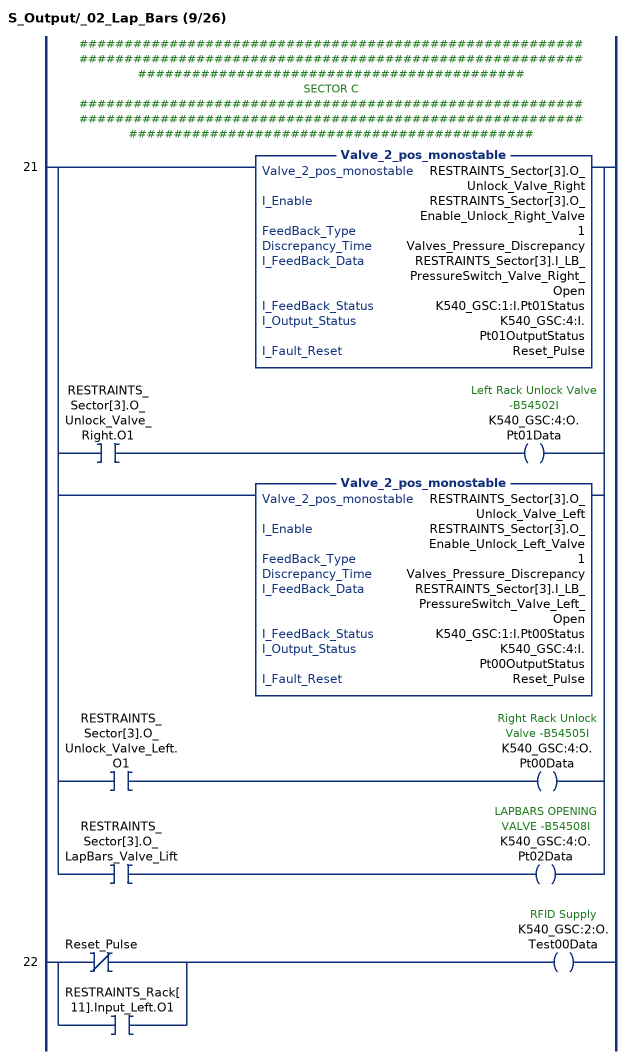
   // ###########################################################################################################################################################
   // SECTOR C
   // #############################################################################################################################################################
   21: [[Valve_2_pos_monostable(RESTRAINTS_Sector[3].O_Unlock_Valve_Right,RESTRAINTS_Sector[3].O_Enable_Unlock_Right_Valve,1,Valves_Pressure_Discrepancy,RESTRAINTS_Sector[3].I_LB_PressureSwitch_Valve_Right_Open,K540_GSC:1:I.Pt01Status,K540_GSC:4:I.Pt01OutputStatus,Reset_Pulse) ,XIC(RESTRAINTS_Sector[3].O_Unlock_Valve_Right.O1) OTE(K540_GSC:4:O.Pt01Data) ] ,[Valve_2_pos_monostable(RESTRAINTS_Sector[3].O_Unlock_Valve_Left,RESTRAINTS_Sector[3].O_Enable_Unlock_Left_Valve,1,Valves_Pressure_Discrepancy,RESTRAINTS_Sector[3].I_LB_PressureSwitch_Valve_Left_Open,K540_GSC:1:I.Pt00Status,K540_GSC:4:I.Pt00OutputStatus,Reset_Pulse) ,XIC(RESTRAINTS_Sector[3].O_Unlock_Valve_Left.O1) OTE(K540_GSC:4:O.Pt00Data) ] ,XIC(RESTRAINTS_Sector[3].O_LapBars_Valve_Lift) OTE(K540_GSC:4:O.Pt02Data) ];
   22: [XIO(Reset_Pulse) ,XIC(RESTRAINTS_Rack[11].Input_Left.O1) ]OTE(K540_GSC:2:O.Test00Data);
